(* CODESYS project Revisora(2)_V3_0_2l.project (continued)
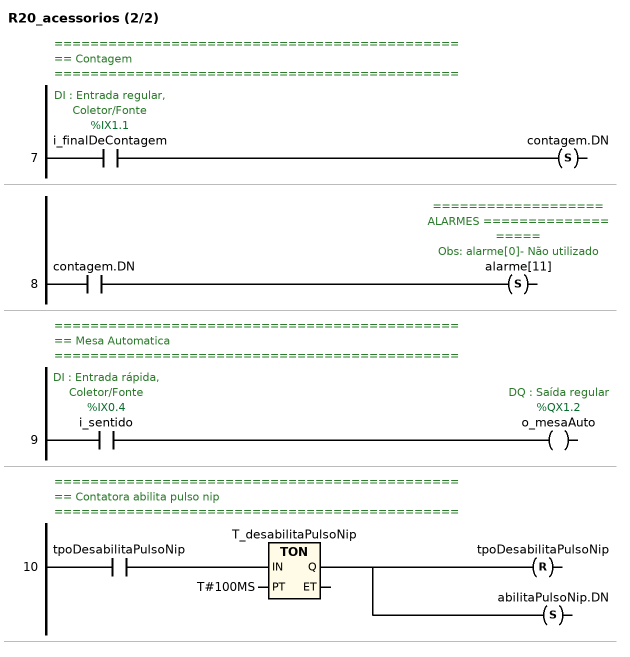
// NETWORK 7
// =============================================
// == Contagem
// =============================================
//   i_finalDeContagem: DI : Entrada regular, Coletor/Fonte | AT %IX1.1
contagem.DN S= i_finalDeContagem;

// NETWORK 8
//   alarme[11]: =================== ALARMES =================== Obs: alarme[0]- Não utilizado
alarme[11] S= contagem.DN;

// NETWORK 9
// =============================================
// == Mesa Automatica
// =============================================
//   i_sentido: DI : Entrada rápida, Coletor/Fonte | AT %IX0.4
//   o_mesaAuto: DQ : Saída regular | AT %QX1.2
o_mesaAuto := i_sentido;

// NETWORK 10
// =============================================
// == Contatora abilita pulso nip
// =============================================
T_desabilitaPulsoNip(IN := tpoDesabilitaPulsoNip, PT := T#100MS); // TON
tpoDesabilitaPulsoNip R= T_desabilitaPulsoNip.Q;
abilitaPulsoNip.DN S= T_desabilitaPulsoNip.Q;

END_PROGRAM

// MyController/Application/01_Maquina/R30_receita
PROGRAM R30_receita
VAR
	
		xtr						: R_TRIG;
		xtf						: F_TRIG;
		atualizaVelocidade		: BOOL;
		tpoVeloc				: TON;
		
		

END_VAR

// Atualização das receitas;
IF triggerBobina THEN
	bobinaAtual.velocDesb:= bobina[numRec].velocDesb;
	//bobinaAtual.torqueDesb:= bobina[1].torqueDesb;
	//bobinaAtual.freioDesb:= bobina[1].freioDesb;
	bobinaAtual.velocReb:= bobina[numRec].velocReb;
	//bobinaAtual.torqueReb:= bobina[1].torqueReb;
	//bobinaAtual.freioReb:= bobina[1].freioReb;
	triggerBobina:= FALSE;
END_IF

// Sentido
IF i_sentido THEN
	sentidoRebobinar:= FALSE;
	sentidoDesbobinar:= TRUE;
	parseAnalog[1]:= bobinaAtual.freioDesb;
	parseAnalog[0]:= bobinaAtual.torqueDesb;
	IF NOT partidaLenta THEN
		M_revisoraVeloc:= bobinaAtual.velocDesb;
	END_IF
ELSE
	sentidoDesbobinar:= FALSE;
	sentidoRebobinar:= TRUE;
	parseAnalog[1]:= bobinaAtual.freioReb;
	parseAnalog[0]:= bobinaAtual.torqueReb;
	IF NOT partidaLenta THEN
		M_revisoraVeloc:= bobinaAtual.velocReb;
	END_IF
END_IF

// Atualização velocidade
xtr(CLK:= i_sentido);
xtf(CLK:= i_sentido);

IF xtr.Q  OR xtf.Q THEN
	atualizaVelocidade:= TRUE;
	//nipMove.IP:= FALSE;
END_IF

//tpoVeloc(IN:= atualizaVelocidade, PT:= T#20MS);

//IF 	tpoVeloc.Q	THEN
//	atualizaVelocidade:= FALSE;
	//IF NOT nipMove.IP THEN
	//		nipMove.IP:= TRUE;
//	END_IF
//END_IF

END_PROGRAM

// MyController/Application/01_Maquina/R50_reset
PROGRAM R50_reset
VAR
END_VAR

IF i_btReset THEN
	
	ihm_alarmeResetInd:= TRUE;
	contagem.DN:= FALSE;
	
ELSE
	
	ihm_alarmeResetInd:= FALSE;
	
END_IF

END_PROGRAM

// MyController/Application/01_Maquina/R99_calcTempos
PROGRAM R99_calcTempos
VAR
END_VAR

// Cálculo dos tempos
tpoInicio:= DINT_TO_TIME(ihm_tempoInicio) * 10;

END_PROGRAM

// MyController/Application/02_Rebobinadores/RB03_analog
PROGRAM RB03_analog
VAR
		calcPorc01				: DINT;
		calcPorc02				: DINT;
END_VAR

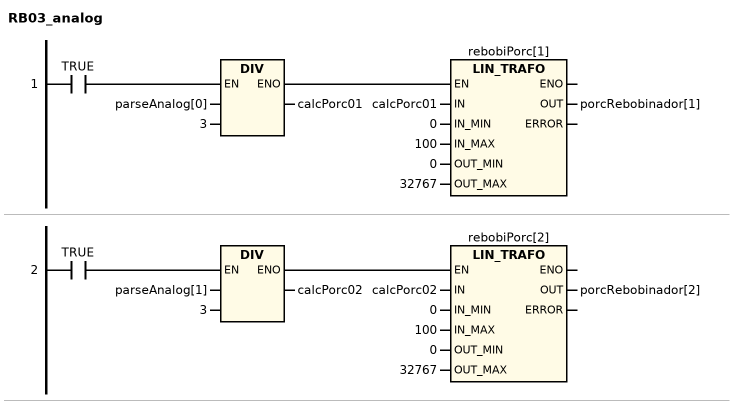
// NETWORK 1
calcPorc01 := parseAnalog[0] / 3;
rebobiPorc[1](
    IN := calcPorc01,
    IN_MIN := 0,
    IN_MAX := 100,
    OUT_MIN := 0,
    OUT_MAX := 32767,
    OUT => porcRebobinador[1]); // LIN_TRAFO

// NETWORK 2
calcPorc02 := parseAnalog[1] / 3;
rebobiPorc[2](
    IN := calcPorc02,
    IN_MIN := 0,
    IN_MAX := 100,
    OUT_MIN := 0,
    OUT_MAX := 32767,
    OUT => porcRebobinador[2]); // LIN_TRAFO

END_PROGRAM

// MyController/Application/02_Rebobinadores/RB04_saidas
PROGRAM RB04_saidas
VAR
END_VAR

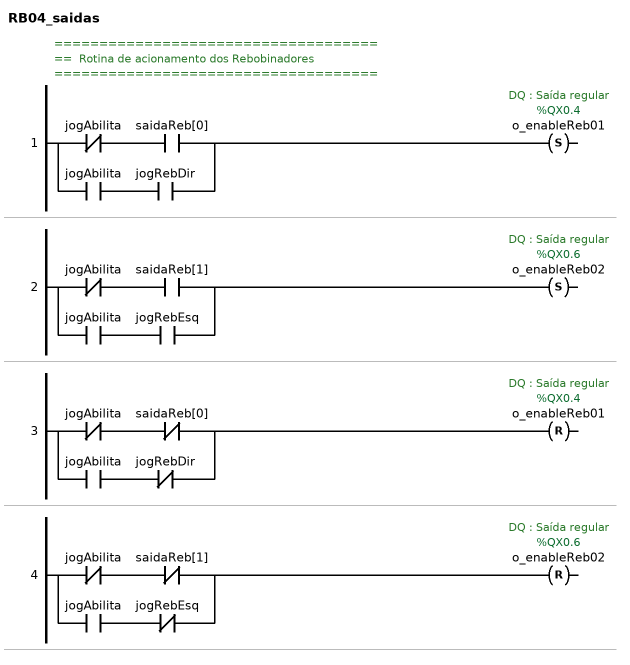
// NETWORK 1
// ====================================
// ==  Rotina de acionamento dos Rebobinadores
// ====================================
//   o_enableReb01: DQ : Saída regular | AT %QX0.4
o_enableReb01 S= NOT jogAbilita AND saidaReb[0] OR jogAbilita AND jogRebDir;

// NETWORK 2
//   o_enableReb02: DQ : Saída regular | AT %QX0.6
o_enableReb02 S= NOT jogAbilita AND saidaReb[1] OR jogAbilita AND jogRebEsq;

// NETWORK 3
//   o_enableReb01: DQ : Saída regular | AT %QX0.4
o_enableReb01 R= NOT jogAbilita AND NOT saidaReb[0] OR jogAbilita AND NOT jogRebDir;

// NETWORK 4
//   o_enableReb02: DQ : Saída regular | AT %QX0.6
o_enableReb02 R= NOT jogAbilita AND NOT saidaReb[1] OR jogAbilita AND NOT jogRebEsq;

END_PROGRAM

// MyController/Application/02_Rebobinadores/RB05_sentido
PROGRAM RB05_sentido
VAR
auxParseAnalog				:ARRAY [1..2] OF REAL;
	T_atrasoTrigger: ARRAY[1..2] OF TON;
	atrasoTrigger: ARRAY[1..2] OF BOOL;
END_VAR

// Calcula quando o valor for menor que 0
//auxParseAnalog[1]:= (parseAnalog[0] * 100) / 1;
//auxParseAnalog[2]:= (parseAnalog[1] * 100) / 1;

T_atrasoTrigger[1](IN := atrasoTrigger[1], PT:= T#200MS); 
T_atrasoTrigger[2](IN := atrasoTrigger[2], PT:= T#200MS);


//atraso para trocar valores
IF triggerValorDesbReb THEN
	atrasoTrigger[1]:=TRUE;
	triggerValorDesbReb:=TRUE;
	IF T_atrasoTrigger[1].Q THEN
		atrasoTrigger[2]:=TRUE;
		M_desbobTorqueOper[1]:=ihm_valorDesb[1];
		M_rebobTorqueOper[1]:=ihm_valorReb[1];
		desbobTorqueOper[1]:=ihm_valorDesb[1];
		rebobTorqueOper[1]:=ihm_valorReb[1];
		M_desbobTorqueOper[2]:=ihm_valorDesb[2];
		M_rebobTorqueOper[2]:=ihm_valorReb[2];
		desbobTorqueOper[2]:=ihm_valorDesb[2];
		rebobTorqueOper[2]:=ihm_valorReb[2];
	END_IF
END_IF
IF  atrasoTrigger[1]= FALSE AND NOT atrasoTrigger[2]= FALSE THEN
		ihm_valorDesb[1]:= desbobTorqueOper[1];
		ihm_valorReb[1]:= rebobTorqueOper[1];
		ihm_valorDesb[2]:= desbobTorqueOper[2];
		ihm_valorReb[2]:= rebobTorqueOper[2];
END_IF
// Reset tempo de atraso
IF T_atrasoTrigger[2].Q THEN
	triggerValorDesbReb:=FALSE;
	atrasoTrigger[1]:= FALSE;
	atrasoTrigger[2]:= FALSE;
END_IF

//auxParseAnalog[1]:=auxAnaloReb01;

IF auxAnaloReb01  + 750 > 10000 THEN
	auxParseAnalog[1]:=10000;
ELSE
	IF i_sentido THEN
		auxParseAnalog[1]:=auxAnaloReb01 + 750;	
	ELSE
		auxParseAnalog[1]:=auxAnaloReb01 ;
	END_IF
END_IF

IF auxAnaloReb02  + 750 > 10000 THEN
	auxParseAnalog[2]:=10000;
ELSE
	IF i_sentido THEN
		auxParseAnalog[2]:=auxAnaloReb02;	
	ELSE
		auxParseAnalog[2]:=auxAnaloReb02  + 750;
	END_IF
END_IF


//IF parseAnalog[0] < 0 THEN
	//valorPorcRebobinador[1]:= auxParseAnalog[1];
//ELSE
	//valorPorcRebobinador[1]:= porcRebobinador[1];	
//END_IF

IF parseAnalog[1] < 0 THEN
	valorPorcRebobinador[2]:= auxParseAnalog[2];
ELSE
	valorPorcRebobinador[2]:= porcRebobinador[2];	
END_IF

// Sentido dos rebobinadores
IF	enbReb.IP THEN
	IF i_sentido THEN
		ladoDir:= FALSE;
		ladoEsq:= TRUE;
		visLadoEsq:= TRUE;
		visLadoDir:= FALSE;
		displayState:= 0;
		valorDesbobTorqueMin:=M_desbobTorqueMin[2];
		valorDesbobTorqueMax:=M_desbobTorqueMax[2];
		valorRebobTorqueMin:=M_rebobTorqueMin[2];
		valorRebobTorqueMax:=M_rebobTorqueMax[2];
	ELSE
		ladoEsq:= FALSE;
		ladoDir:= TRUE;
		visLadoEsq:= FALSE;
		visLadoDir:= TRUE;
		displayState:= 1;
		
		valorRebobTorqueMin:=M_desbobTorqueMin[1];
		valorRebobTorqueMax:=M_desbobTorqueMax[1];
		valorDesbobTorqueMin:=M_rebobTorqueMin[1];
		valorDesbobTorqueMax:=M_rebobTorqueMax[1];
	END_IF
END_IF

// Editar valores

IF ligaMaq THEN
	IF ladoEsq THEN
		analoReb02:= REAL_TO_INT((auxParseAnalog[1])*-1); 
		analoReb01:= REAL_TO_INT((auxParseAnalog[2]));
		delayTorq[0] := T#500MS;
		delayTorq[1] := T#0MS;
		
	END_IF
	
	IF ladoDir THEN
		analoReb02:= REAL_TO_INT(auxParseAnalog[2])*-1;
		analoReb01:= REAL_TO_INT(auxParseAnalog[1]);
		delayTorq[0] := T#0MS;
		delayTorq[1] := T#500MS;
	END_IF
END_IF
	//IF NOT ciclo.IP THEN
	//	ladoEsq:= FALSE;
	//	ladoDir:= FALSE;
//	END_IF
	
	// Parada
	IF torqueParada THEN
		IF ladoEsq THEN
			analoReb02:= 3000;
			analoReb01:= 3000;
		ELSE
			analoReb02:= -3000;
			analoReb01:= -3000;
		END_IF
	END_IF
// Calcula quando o valor for menor que 0
//auxParseAnalog[1]:= (parseAnalog[0] * 328) / 3;
//auxParseAnalog[2]:= (parseAnalog[1] * 328) / 3;

END_PROGRAM

// MyController/Application/03_Nip/NP01_geral
PROGRAM NP01_geral
VAR
	TD_power				: TOF;
END_VAR
VAR // added by the converter: edge detectors and wires of the graphical bodies
    _ft1 : F_TRIG;
END_VAR

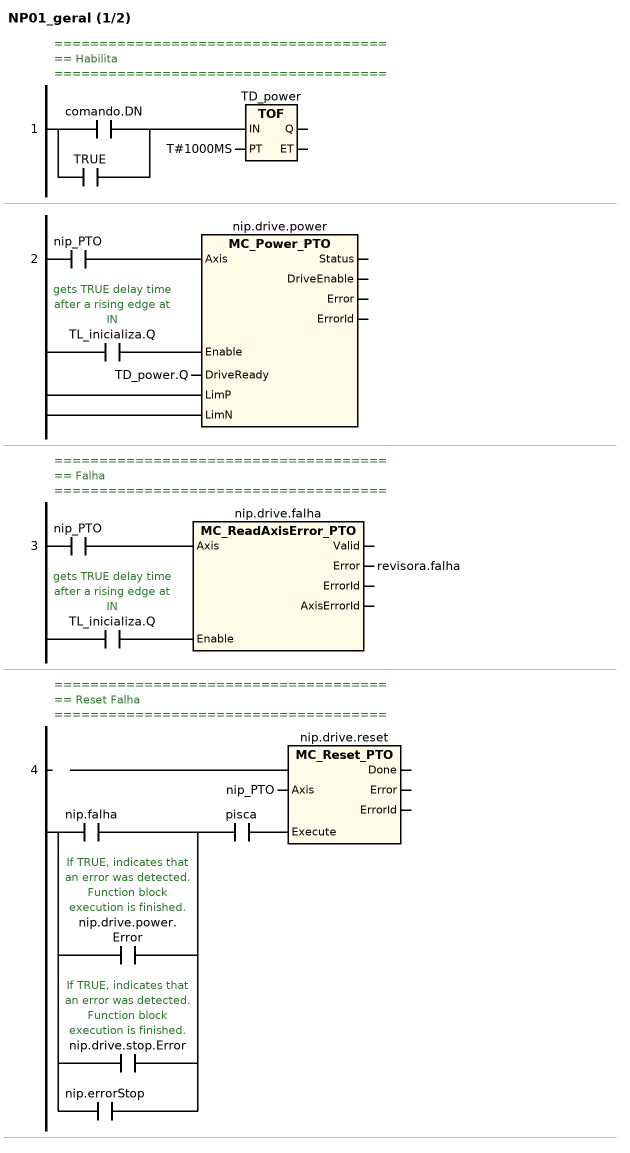
// NETWORK 1
// =====================================
// == Habilita
// =====================================
TD_power(IN := comando.DN OR TRUE, PT := T#1000MS); // TOF

// NETWORK 2
//   TL_inicializa.Q: gets TRUE delay time after a rising edge at IN
//   TD_power.Q: gets FALSE, when PT milliseconds elapsed, since falling edge at IN
nip.drive.power(
    Axis := nip_PTO,
    Enable := TL_inicializa.Q,
    DriveReady := TD_power.Q,
    LimP := TRUE,
    LimN := TRUE); // MC_Power_PTO

// NETWORK 3
// =====================================
// == Falha
// =====================================
//   TL_inicializa.Q: gets TRUE delay time after a rising edge at IN
nip.drive.falha(Axis := nip_PTO, Enable := TL_inicializa.Q, Error => revisora.falha); // MC_ReadAxisError_PTO

// NETWORK 4
// =====================================
// == Reset Falha
// =====================================
//   nip.drive.power.Error: If TRUE, indicates that an error was detected. Function block execution is finished.
//   nip.drive.stop.Error: If TRUE, indicates that an error was detected. Function block execution is finished.
nip.drive.reset(Axis := nip_PTO, Execute := (nip.falha OR nip.drive.power.Error OR nip.drive.stop.Error OR nip.errorStop) AND pisca); // MC_Reset_PTO

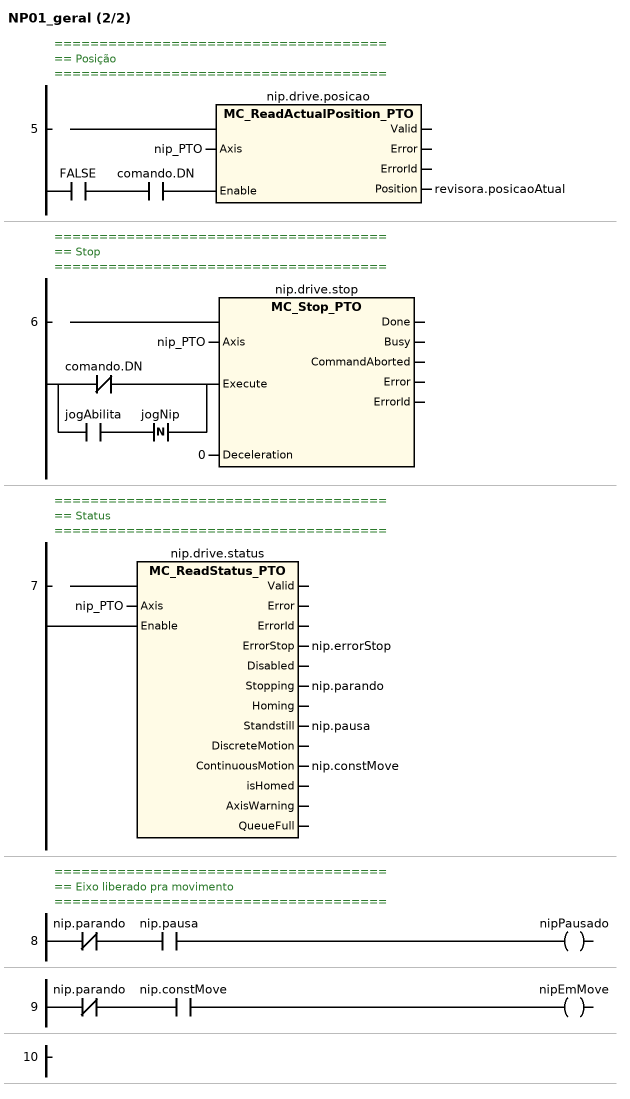
// NETWORK 5
// =====================================
// == Posição
// =====================================
nip.drive.posicao(Axis := nip_PTO, Enable := FALSE AND comando.DN, Position => revisora.posicaoAtual); // MC_ReadActualPosition_PTO

// NETWORK 6
// =====================================
// == Stop
// =====================================
_ft1(CLK := jogNip);
nip.drive.stop(Axis := nip_PTO, Execute := NOT comando.DN OR jogAbilita AND _ft1.Q, Deceleration := 0); // MC_Stop_PTO

// NETWORK 7
// =====================================
// == Status
// =====================================
nip.drive.status(
    Axis := nip_PTO,
    Enable := TRUE,
    ErrorStop => nip.errorStop,
    Stopping => nip.parando,
    Standstill => nip.pausa,
    ContinuousMotion => nip.constMove); // MC_ReadStatus_PTO

// NETWORK 8
// =====================================
// == Eixo liberado pra movimento
// =====================================
nipPausado := NOT nip.parando AND nip.pausa;

// NETWORK 9
nipEmMove := NOT nip.parando AND nip.constMove;

// NETWORK 10

END_PROGRAM

// MyController/Application/03_Nip/NP02_enableNip
PROGRAM NP02_enableNip
VAR
END_VAR
VAR // added by the converter: edge detectors and wires of the graphical bodies
    _ft1 : F_TRIG;
END_VAR

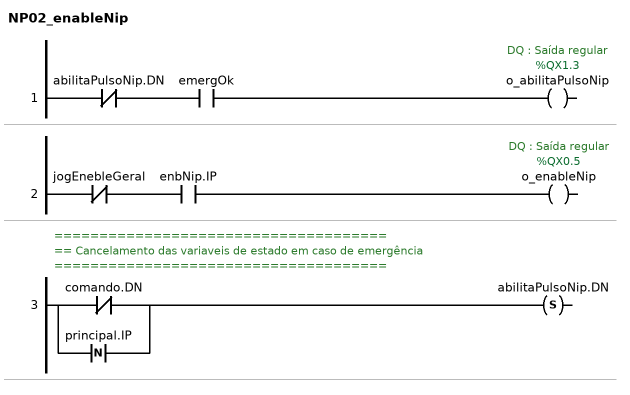
// NETWORK 1
//   o_abilitaPulsoNip: DQ : Saída regular | AT %QX1.3
o_abilitaPulsoNip := NOT abilitaPulsoNip.DN AND emergOk;

// NETWORK 2
//   o_enableNip: DQ : Saída regular | AT %QX0.5
o_enableNip := NOT jogEnebleGeral AND enbNip.IP;

// NETWORK 3
// =====================================
// == Cancelamento das variaveis de estado em caso de emergência
// =====================================
_ft1(CLK := principal.IP);
abilitaPulsoNip.DN S= NOT comando.DN OR _ft1.Q;

END_PROGRAM

// MyController/Application/03_Nip/NP03_auto
PROGRAM NP03_auto
VAR
	TF_enable						: TON;
END_VAR
VAR // added by the converter: edge detectors and wires of the graphical bodies
    _rt1, _rt2 : R_TRIG;
    _w1, _w2 : BOOL;
    _ft1 : F_TRIG;
END_VAR

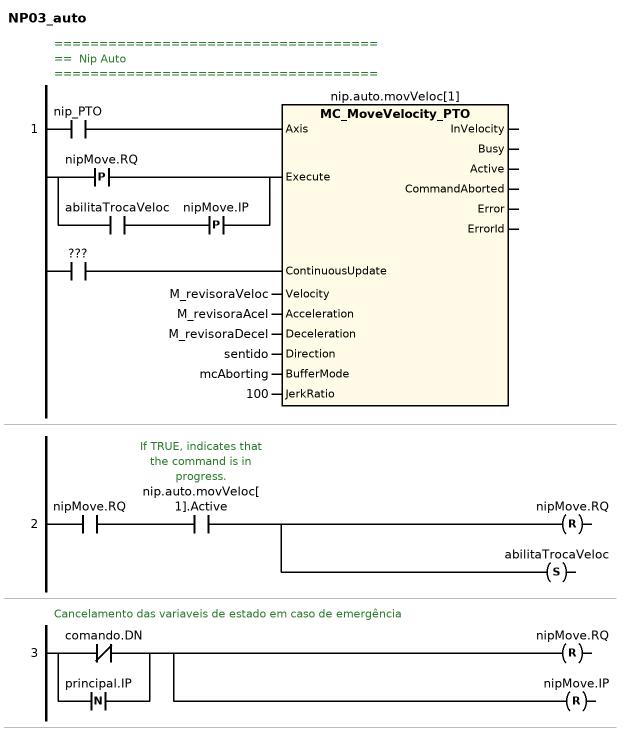
// NETWORK 1
// ====================================
// ==  Nip Auto
// ====================================
_rt1(CLK := nipMove.RQ);
_rt2(CLK := nipMove.IP);
nip.auto.movVeloc[1](
    Axis := nip_PTO,
    Execute := _rt1.Q OR abilitaTrocaVeloc AND _rt2.Q,
    Velocity := M_revisoraVeloc,
    Acceleration := M_revisoraAcel,
    Deceleration := M_revisoraDecel,
    Direction := sentido,
    BufferMode := mcAborting,
    JerkRatio := 100); // MC_MoveVelocity_PTO

// NETWORK 2
//   nip.auto.movVeloc[1].Active: If TRUE, indicates that the command is in progress.
_w1 := nipMove.RQ AND nip.auto.movVeloc[1].Active;
nipMove.RQ R= _w1;
abilitaTrocaVeloc S= _w1;

// NETWORK 3
// Cancelamento das variaveis de estado em caso de emergência
_ft1(CLK := principal.IP);
_w2 := NOT comando.DN OR _ft1.Q;
nipMove.RQ R= _w2;
nipMove.IP R= _w2;

END_PROGRAM

// MyController/Application/03_Nip/NP04_parada
PROGRAM NP04_parada
VAR
	
	job: BOOL;
	T_DelayPosVeloc: TON;
	T_atraso: TON;
END_VAR
VAR // added by the converter: edge detectors and wires of the graphical bodies
    _rt1 : R_TRIG;
    _w1, _w2 : BOOL;
    _ft1 : F_TRIG;
END_VAR

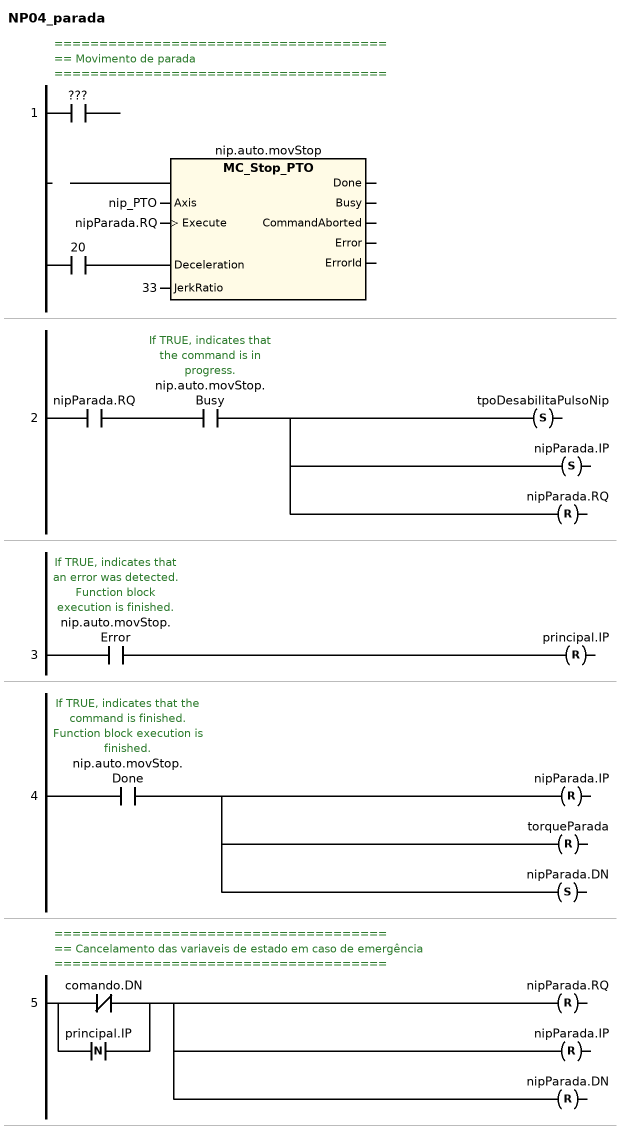
// NETWORK 1
// =====================================
// == Movimento de parada
// =====================================
_rt1(CLK := nipParada.RQ);
nip.auto.movStop(Axis := nip_PTO, Execute := _rt1.Q, Deceleration := 20, JerkRatio := 33); // MC_Stop_PTO

// NETWORK 2
//   nip.auto.movStop.Busy: If TRUE, indicates that the command is in progress.
_w1 := nipParada.RQ AND nip.auto.movStop.Busy;
tpoDesabilitaPulsoNip S= _w1;
nipParada.IP S= _w1;
nipParada.RQ R= _w1;

// NETWORK 3
//   nip.auto.movStop.Error: If TRUE, indicates that an error was detected. Function block execution is finished.
principal.IP R= nip.auto.movStop.Error;

// NETWORK 4
//   nip.auto.movStop.Done: If TRUE, indicates that the command is finished. Function block execution is finished.
nipParada.IP R= nip.auto.movStop.Done;
torqueParada R= nip.auto.movStop.Done;
nipParada.DN S= nip.auto.movStop.Done;

// NETWORK 5
// =====================================
// == Cancelamento das variaveis de estado em caso de emergência
// =====================================
_ft1(CLK := principal.IP);
_w2 := NOT comando.DN OR _ft1.Q;
nipParada.RQ R= _w2;
nipParada.IP R= _w2;
nipParada.DN R= _w2;

END_PROGRAM

// MyController/Application/03_Nip/NP06_jog
PROGRAM NP06_jog
VAR
	auxJogPos								: BOOL;
	auxJopNeg								: BOOL;
END_VAR
VAR // added by the converter: edge detectors and wires of the graphical bodies
    _ft1, _ft2 : F_TRIG;
END_VAR

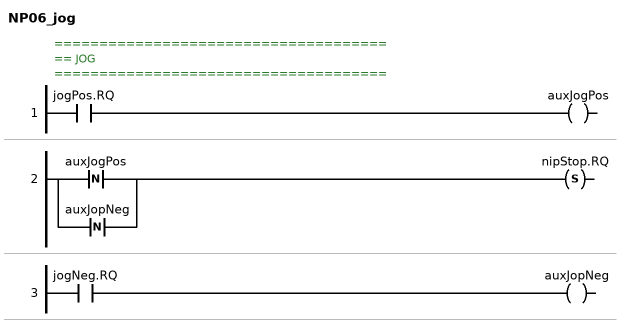
// NETWORK 1
// =====================================
// == JOG
// =====================================
auxJogPos := jogPos.RQ;

// NETWORK 2
_ft1(CLK := auxJogPos);
_ft2(CLK := auxJopNeg);
nipStop.RQ S= _ft1.Q OR _ft2.Q;

// NETWORK 3
auxJopNeg := jogNeg.RQ;

END_PROGRAM

// MyController/Application/03_Nip/NP07_veloc
PROGRAM NP07_veloc
VAR

	timerVeloc 		: TON;

END_VAR

// Partida Lenta


IF sentido = -1 THEN
	M_revisoraVeloc:=(bobinaAtual.velocReb );
END_IF
IF sentido = 1 THEN
	M_revisoraVeloc:=(bobinaAtual.velocDesb );
END_IF

//IF nipMove.RQ THEN
//	IF bobinaAtual.velocDesb > 800 OR bobinaAtual.velocReb > 800 THEN	
	//	M_revisoraVeloc:= 600;
	//	partidaLenta:= TRUE;
//	END_IF
//END_IF

//timerVeloc(IN:= partidaLenta, PT:= T#7S);

//IF 	timerVeloc.Q THEN
	//nipMove.IP:= FALSE;
	//partidaLenta:= FALSE;
	//IF i_sentido THEN
	//	M_revisoraVeloc:= bobinaAtual.velocDesb;
	//	nipMove.IP:= TRUE;
//	ELSE
//		M_revisoraVeloc:= bobinaAtual.velocReb;
//		nipMove.IP:= TRUE;
//	END_IF
//END_IF

//IF NOT comando.DN OR principal.IP OR ligaMaq THEN
//	partidaLenta:= FALSE;
//END_IF

END_PROGRAM

// MyController/Application/03_Nip/NP09_sentido
PROGRAM NP09_sentido
VAR
END_VAR

// Mudança de sentido
IF i_sentido AND NOT ciclo.IP THEN
	sentido:= 1;
	M_pulsosParar:= 20;
ELSIF NOT i_sentido AND NOT ciclo.IP THEN
	sentido:= -1;
	M_pulsosParar:= -20;
END_IF

END_PROGRAM

// MyController/Application/03_Nip/NP20_JogTest
PROGRAM NP20_JogTest
VAR
	auxVeloc			:DINT;
	auxReb01			: INT;
	auxReb02			: INT;
END_VAR

IF jogVelocNip >3000 THEN
	jogVelocNip:= 3000;
	
END_IF

IF jogAbilita = TRUE THEN
	revisoraVelocNip:=jogVelocNip;
ELSE
	revisoraVelocNip:=M_revisoraVeloc;
END_IF

END_PROGRAM

// MyController/Application/19_Ultra/U10_auto
PROGRAM U10_auto
VAR
	auxBit						: BOOL;
	auxReal						: REAL;
	auxTorque					: ARRAY[0..4] OF REAL;
	desbobEscalaTorque			: ARRAY[0..4] OF LIN_TRAFO;
	rebobEscalaTorque			: ARRAY[0..4] OF LIN_TRAFO;
	rebobTorqueRamp				: DINT:= 200;
	sinalUltraSom				: ARRAY[1..2] OF INT;
	TL_rebobOk					: TON;
	ultraSomEscala				: LIN_TRAFO;
	porcUltraSom				: ARRAY[1..2] OF REAL;
	desbobEscalaUltraSom		: ARRAY[0..4] OF LIN_TRAFO;
	rebobEscalaUltraSom			: ARRAY[0..4] OF LIN_TRAFO;
END_VAR
VAR // added by the converter: edge detectors and wires of the graphical bodies
    _rt1, _rt2, _rt3, _rt4 : R_TRIG;
    _w1, _w2, _w3, _w4, _w5, _w6, _w7, _w8, _w9, _w10, _w11, _w12 : BOOL;
END_VAR

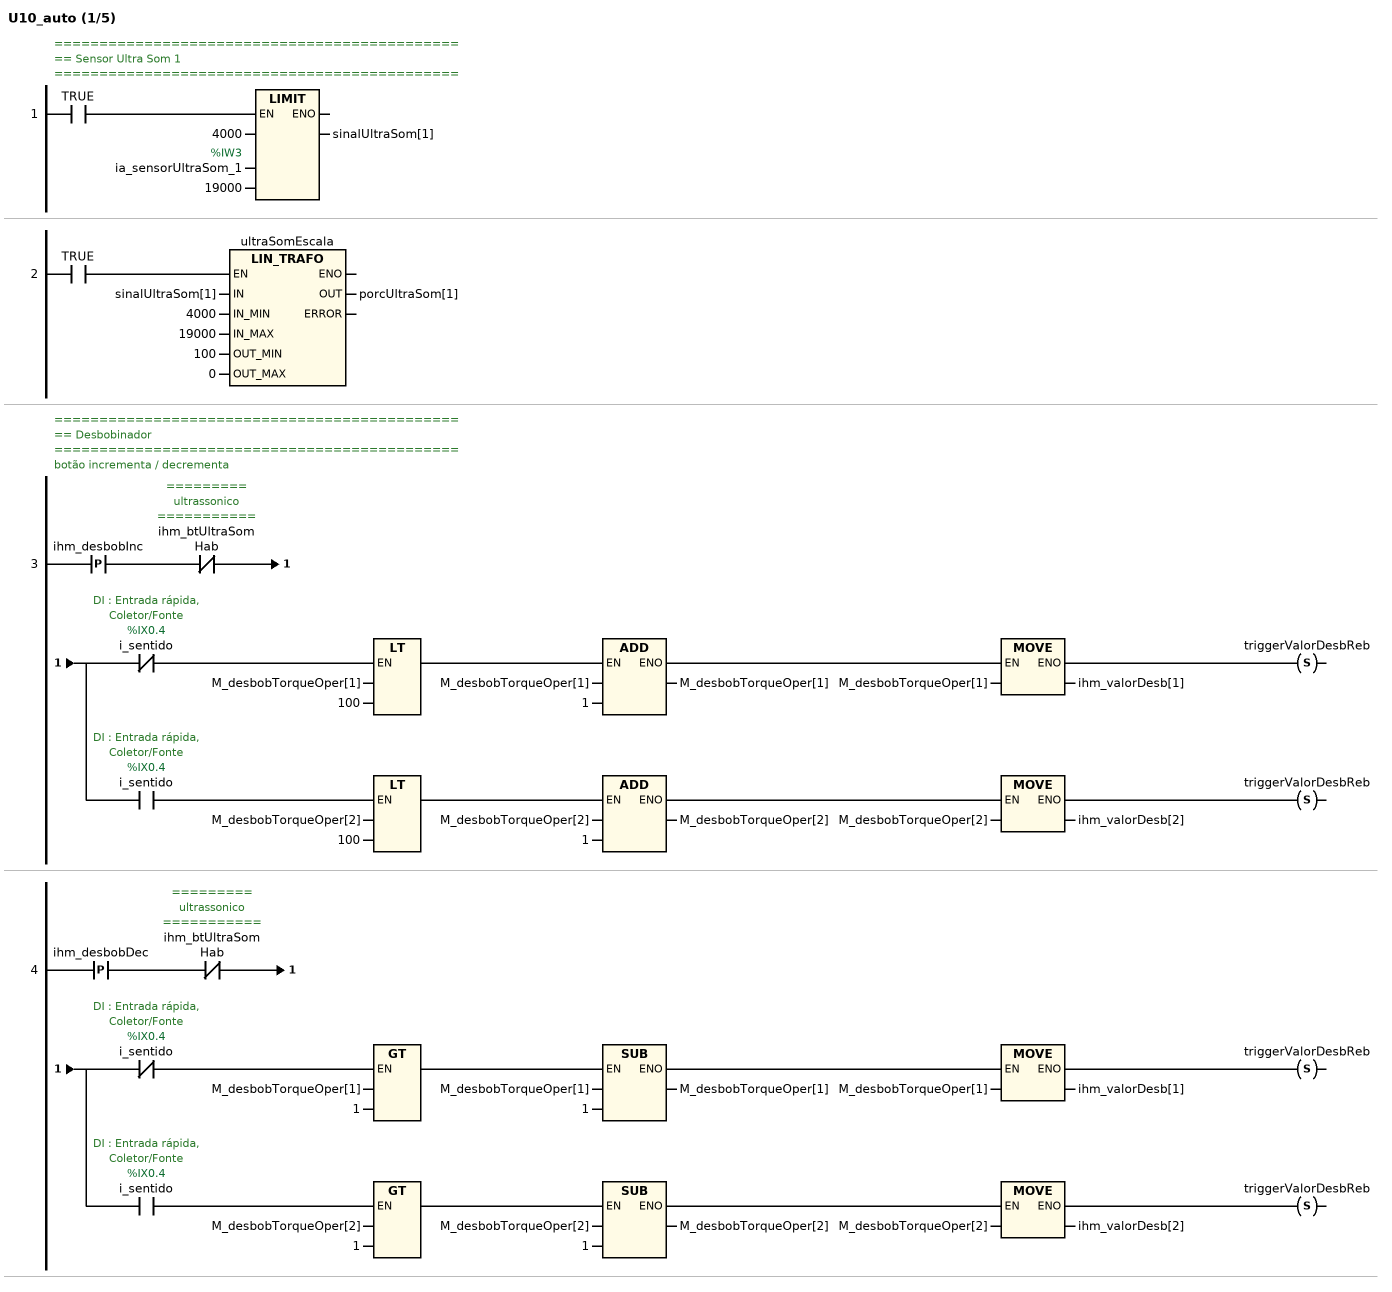
// NETWORK 1
// =============================================
// == Sensor Ultra Som 1
// =============================================
//   ia_sensorUltraSom_1: Entradas_Analog : | AT %IW3
sinalUltraSom[1] := LIMIT(4000, ia_sensorUltraSom_1, 19000);

// NETWORK 2
ultraSomEscala(
    IN := sinalUltraSom[1],
    IN_MIN := 4000,
    IN_MAX := 19000,
    OUT_MIN := 100,
    OUT_MAX := 0,
    OUT => porcUltraSom[1]); // LIN_TRAFO

// NETWORK 3
// =============================================
// == Desbobinador
// =============================================
// botão incrementa / decrementa
//   ihm_btUltraSomHab: ========= ultrassonico ===========
//   i_sentido: DI : Entrada rápida, Coletor/Fonte | AT %IX0.4
_rt1(CLK := ihm_desbobInc);
_w1 := _rt1.Q AND NOT ihm_btUltraSomHab;
IF _w1 AND NOT i_sentido AND M_desbobTorqueOper[1] < 100 THEN
    M_desbobTorqueOper[1] := M_desbobTorqueOper[1] + 1;
END_IF
IF _w1 AND NOT i_sentido AND M_desbobTorqueOper[1] < 100 THEN ihm_valorDesb[1] := M_desbobTorqueOper[1]; END_IF
triggerValorDesbReb S= _w1 AND NOT i_sentido AND M_desbobTorqueOper[1] < 100;
IF _w1 AND i_sentido AND M_desbobTorqueOper[2] < 100 THEN
    M_desbobTorqueOper[2] := M_desbobTorqueOper[2] + 1;
END_IF
IF _w1 AND i_sentido AND M_desbobTorqueOper[2] < 100 THEN ihm_valorDesb[2] := M_desbobTorqueOper[2]; END_IF
triggerValorDesbReb S= _w1 AND i_sentido AND M_desbobTorqueOper[2] < 100;

// NETWORK 4
//   ihm_btUltraSomHab: ========= ultrassonico ===========
//   i_sentido: DI : Entrada rápida, Coletor/Fonte | AT %IX0.4
_rt2(CLK := ihm_desbobDec);
_w2 := _rt2.Q AND NOT ihm_btUltraSomHab;
IF _w2 AND NOT i_sentido AND M_desbobTorqueOper[1] > 1 THEN
    M_desbobTorqueOper[1] := M_desbobTorqueOper[1] - 1;
END_IF
IF _w2 AND NOT i_sentido AND M_desbobTorqueOper[1] > 1 THEN ihm_valorDesb[1] := M_desbobTorqueOper[1]; END_IF
triggerValorDesbReb S= _w2 AND NOT i_sentido AND M_desbobTorqueOper[1] > 1;
IF _w2 AND i_sentido AND M_desbobTorqueOper[2] > 1 THEN M_desbobTorqueOper[2] := M_desbobTorqueOper[2] - 1; END_IF
IF _w2 AND i_sentido AND M_desbobTorqueOper[2] > 1 THEN ihm_valorDesb[2] := M_desbobTorqueOper[2]; END_IF
triggerValorDesbReb S= _w2 AND i_sentido AND M_desbobTorqueOper[2] > 1;

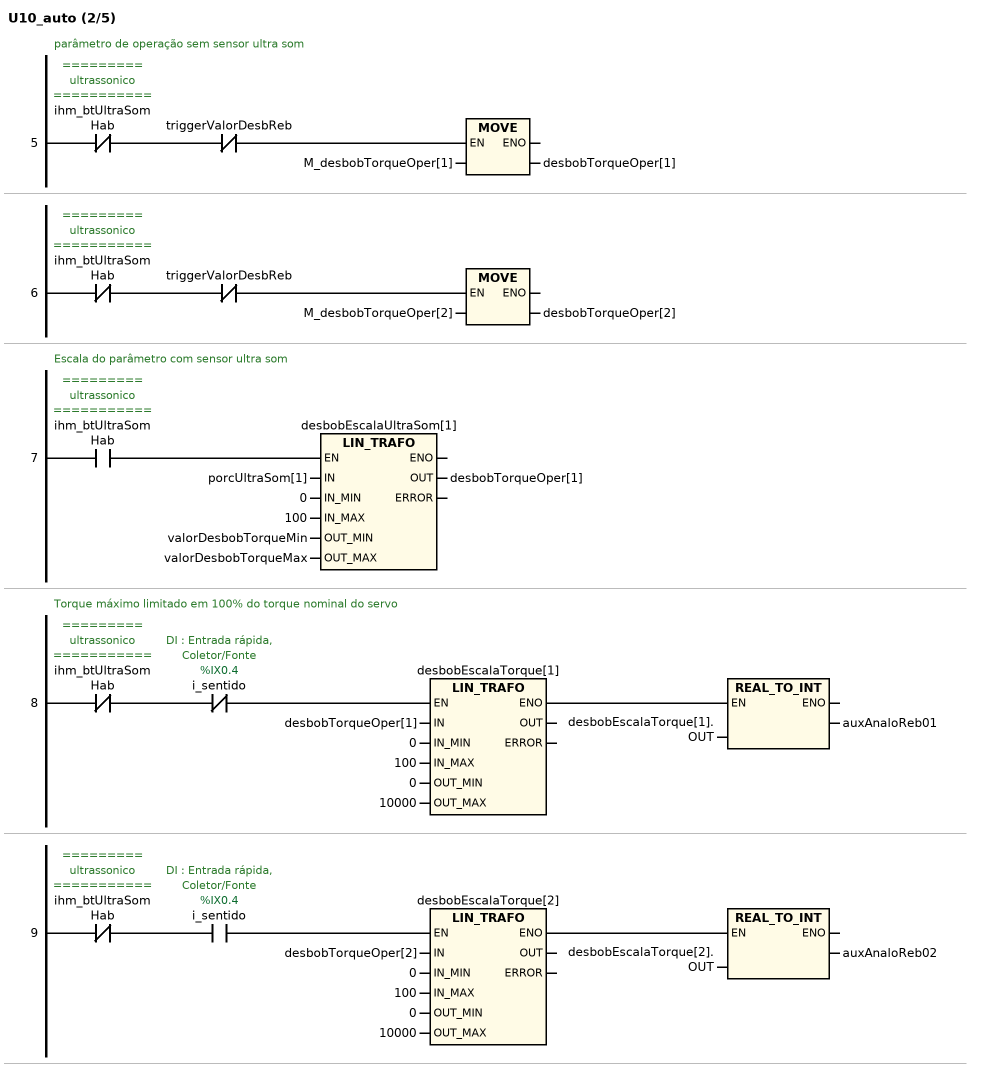
// NETWORK 5
// parâmetro de operação sem sensor ultra som
//   ihm_btUltraSomHab: ========= ultrassonico ===========
IF NOT ihm_btUltraSomHab AND NOT triggerValorDesbReb THEN desbobTorqueOper[1] := M_desbobTorqueOper[1]; END_IF

// NETWORK 6
//   ihm_btUltraSomHab: ========= ultrassonico ===========
IF NOT ihm_btUltraSomHab AND NOT triggerValorDesbReb THEN desbobTorqueOper[2] := M_desbobTorqueOper[2]; END_IF

// NETWORK 7
// Escala do parâmetro com sensor ultra som
//   ihm_btUltraSomHab: ========= ultrassonico ===========
IF ihm_btUltraSomHab THEN
    desbobEscalaUltraSom[1](
        IN := porcUltraSom[1],
        IN_MIN := 0,
        IN_MAX := 100,
        OUT_MIN := valorDesbobTorqueMin,
        OUT_MAX := valorDesbobTorqueMax,
        OUT => desbobTorqueOper[1]); // LIN_TRAFO
END_IF

// NETWORK 8
// Torque máximo limitado em 100% do torque nominal do servo
//   ihm_btUltraSomHab: ========= ultrassonico ===========
//   i_sentido: DI : Entrada rápida, Coletor/Fonte | AT %IX0.4
//   desbobEscalaTorque[1].OUT: output value
_w3 := NOT ihm_btUltraSomHab AND NOT i_sentido;
IF _w3 THEN
    desbobEscalaTorque[1](IN := desbobTorqueOper[1], IN_MIN := 0, IN_MAX := 100, OUT_MIN := 0, OUT_MAX := 10000); // LIN_TRAFO
END_IF
IF _w3 THEN auxAnaloReb01 := REAL_TO_INT(desbobEscalaTorque[1].OUT); END_IF

// NETWORK 9
//   ihm_btUltraSomHab: ========= ultrassonico ===========
//   i_sentido: DI : Entrada rápida, Coletor/Fonte | AT %IX0.4
//   desbobEscalaTorque[2].OUT: output value
_w4 := NOT ihm_btUltraSomHab AND i_sentido;
IF _w4 THEN
    desbobEscalaTorque[2](IN := desbobTorqueOper[2], IN_MIN := 0, IN_MAX := 100, OUT_MIN := 0, OUT_MAX := 10000); // LIN_TRAFO
END_IF
IF _w4 THEN auxAnaloReb02 := REAL_TO_INT(desbobEscalaTorque[2].OUT); END_IF

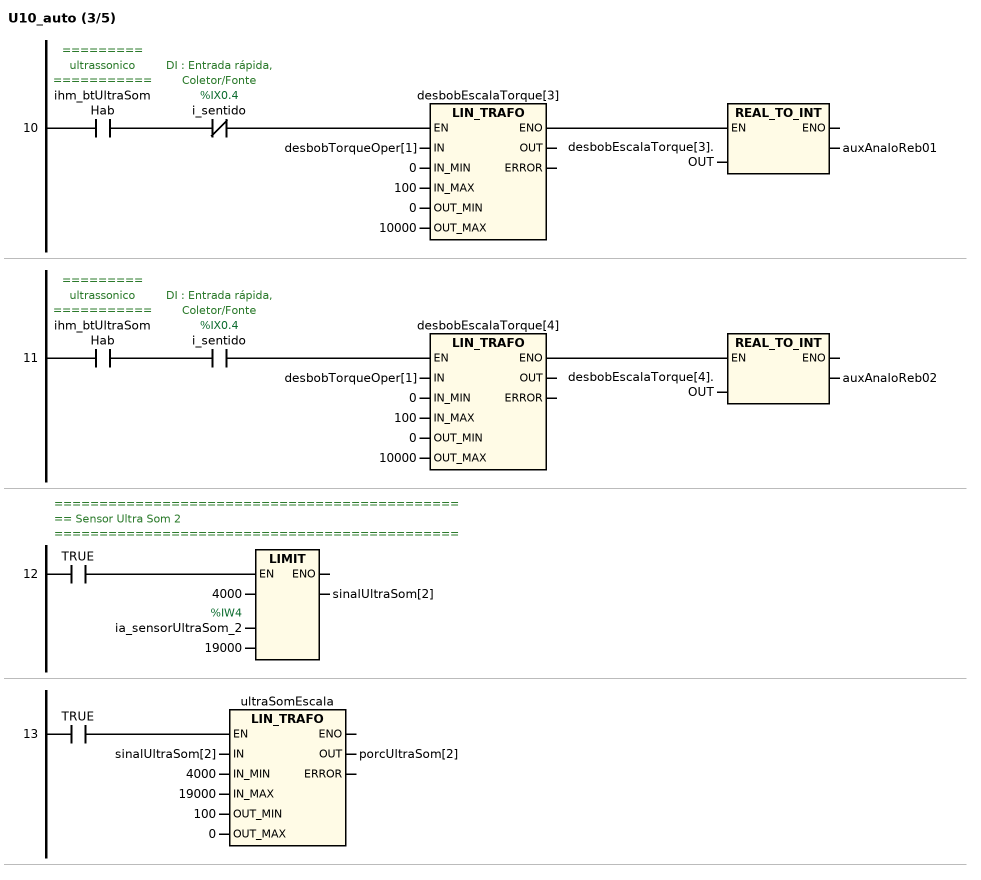
// NETWORK 10
//   ihm_btUltraSomHab: ========= ultrassonico ===========
//   i_sentido: DI : Entrada rápida, Coletor/Fonte | AT %IX0.4
//   desbobEscalaTorque[3].OUT: output value
_w5 := ihm_btUltraSomHab AND NOT i_sentido;
IF _w5 THEN
    desbobEscalaTorque[3](IN := desbobTorqueOper[1], IN_MIN := 0, IN_MAX := 100, OUT_MIN := 0, OUT_MAX := 10000); // LIN_TRAFO
END_IF
IF _w5 THEN auxAnaloReb01 := REAL_TO_INT(desbobEscalaTorque[3].OUT); END_IF

// NETWORK 11
//   ihm_btUltraSomHab: ========= ultrassonico ===========
//   i_sentido: DI : Entrada rápida, Coletor/Fonte | AT %IX0.4
//   desbobEscalaTorque[4].OUT: output value
_w6 := ihm_btUltraSomHab AND i_sentido;
IF _w6 THEN
    desbobEscalaTorque[4](IN := desbobTorqueOper[1], IN_MIN := 0, IN_MAX := 100, OUT_MIN := 0, OUT_MAX := 10000); // LIN_TRAFO
END_IF
IF _w6 THEN auxAnaloReb02 := REAL_TO_INT(desbobEscalaTorque[4].OUT); END_IF

// NETWORK 12
// =============================================
// == Sensor Ultra Som 2
// =============================================
//   ia_sensorUltraSom_2: Entradas_Analog : | AT %IW4
sinalUltraSom[2] := LIMIT(4000, ia_sensorUltraSom_2, 19000);

// NETWORK 13
ultraSomEscala(
    IN := sinalUltraSom[2],
    IN_MIN := 4000,
    IN_MAX := 19000,
    OUT_MIN := 100,
    OUT_MAX := 0,
    OUT => porcUltraSom[2]); // LIN_TRAFO

